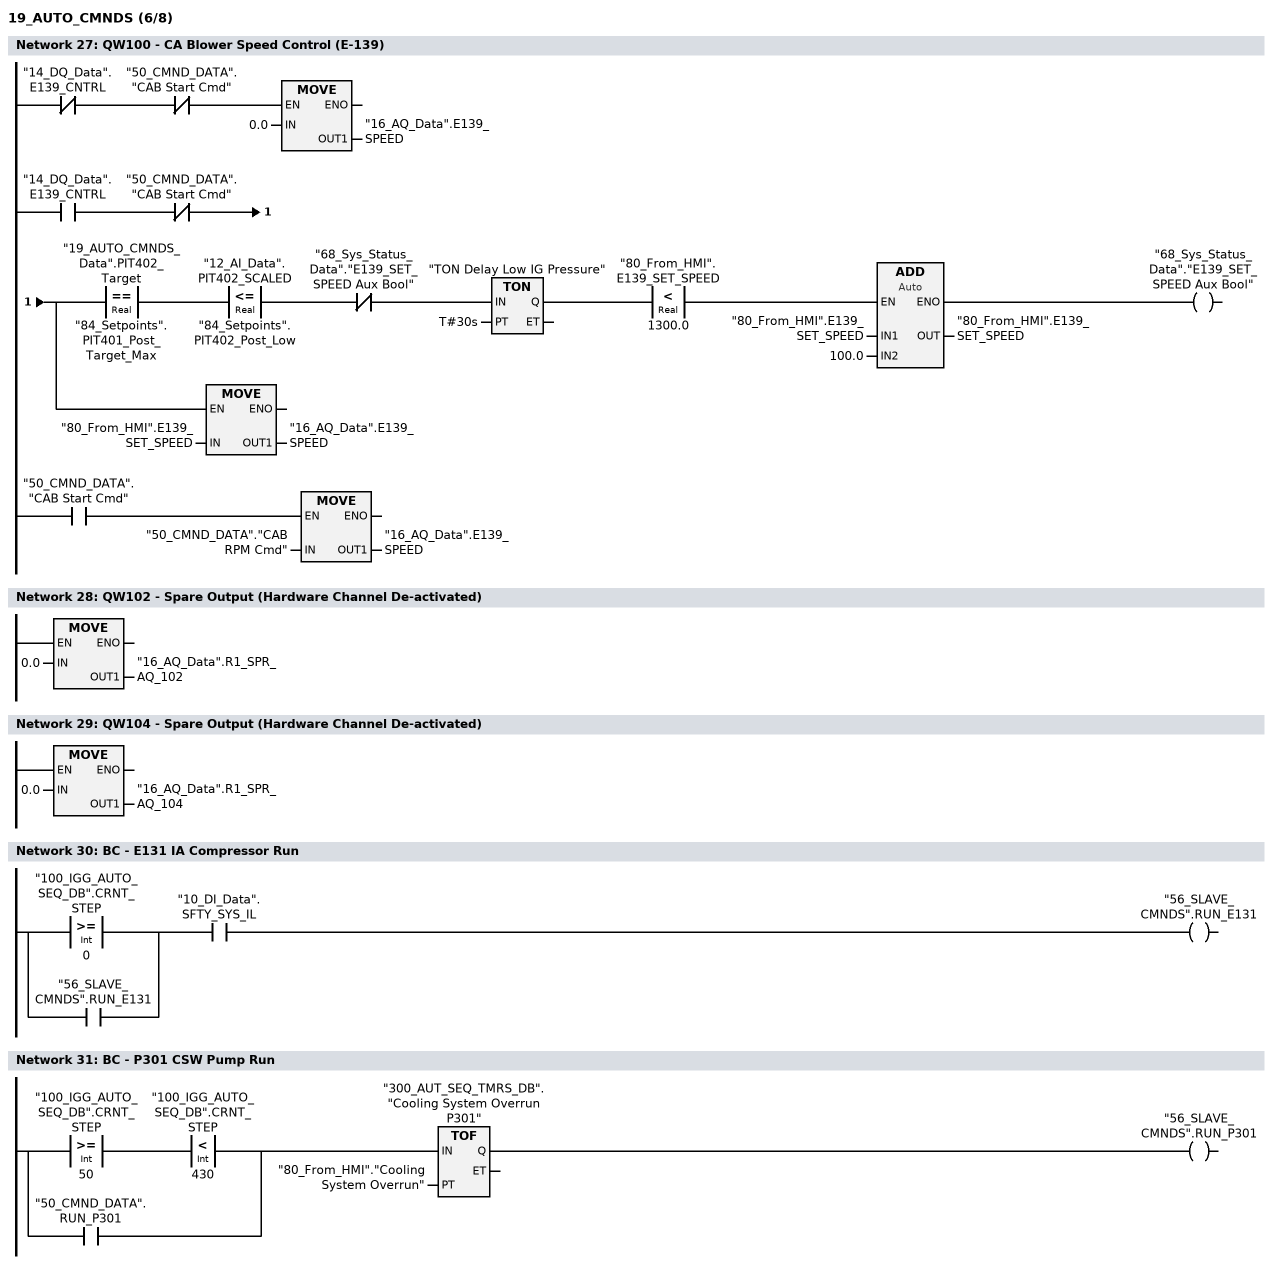
   IF NOT "14_DQ_Data".E139_CNTRL AND NOT "50_CMND_DATA"."CAB Start Cmd" THEN
       "16_AQ_Data".E139_SPEED := 0.0;
   END_IF;
   #_w1 := "14_DQ_Data".E139_CNTRL AND NOT "50_CMND_DATA"."CAB Start Cmd";
   "TON Delay Low IG Pressure".TON(IN := #_w1 AND ("19_AUTO_CMNDS_Data".PIT402_Target = "84_Setpoints".PIT401_Post_Target_Max) AND ("12_AI_Data".PIT402_SCALED <= "84_Setpoints".PIT402_Post_Low) AND NOT "68_Sys_Status_Data"."E139_SET_SPEED Aux Bool",
                           PT := T#30s);
   #_w2 := "TON Delay Low IG Pressure".Q AND ("80_From_HMI".E139_SET_SPEED < 1300.0);
   IF #_w2 THEN "80_From_HMI".E139_SET_SPEED := "80_From_HMI".E139_SET_SPEED + 100.0; END_IF;
   "68_Sys_Status_Data"."E139_SET_SPEED Aux Bool" := #_w2;
   IF #_w1 THEN "16_AQ_Data".E139_SPEED := "80_From_HMI".E139_SET_SPEED; END_IF;
   IF "50_CMND_DATA"."CAB Start Cmd" THEN "16_AQ_Data".E139_SPEED := "50_CMND_DATA"."CAB RPM Cmd"; END_IF;
END_REGION

REGION Network 28: QW102 - Spare Output (Hardware Channel De-activated)
   RUNG wire#powerrail
      Move(in := 0.0, out1 => "16_AQ_Data".R1_SPR_AQ_102)
   END_RUNG
   // the same network as SCL:
   "16_AQ_Data".R1_SPR_AQ_102 := 0.0;
END_REGION

REGION Network 29: QW104 - Spare Output (Hardware Channel De-activated)
   RUNG wire#powerrail
      Move(in := 0.0, out1 => "16_AQ_Data".R1_SPR_AQ_104)
   END_RUNG
   // the same network as SCL:
   "16_AQ_Data".R1_SPR_AQ_104 := 0.0;
END_REGION

REGION Network 30: BC - E131 IA Compressor Run
   RUNG wire#powerrail
      { S7_Templates := "SrcType := Int" } GE_Contact(in1 := "100_IGG_AUTO_SEQ_DB".CRNT_STEP, in2 := 0)
      wire#w1
      Contact( "10_DI_Data".SFTY_SYS_IL )
      Coil( "56_SLAVE_CMNDS".RUN_E131 )
   END_RUNG
   RUNG wire#powerrail
      Contact( "56_SLAVE_CMNDS".RUN_E131 )
   END_RUNG wire#w1
   // the same network as SCL:
   "56_SLAVE_CMNDS".RUN_E131 := (("100_IGG_AUTO_SEQ_DB".CRNT_STEP >= 0) OR "56_SLAVE_CMNDS".RUN_E131) AND "10_DI_Data".SFTY_SYS_IL;
END_REGION

REGION Network 31: BC - P301 CSW Pump Run
   "300_AUT_SEQ_TMRS_DB"."Cooling System Overrun P301".TOF(IN := (("100_IGG_AUTO_SEQ_DB".CRNT_STEP >= 50) AND ("100_IGG_AUTO_SEQ_DB".CRNT_STEP < 430)) OR "50_CMND_DATA".RUN_P301,
                           PT := "80_From_HMI"."Cooling System Overrun");
   "56_SLAVE_CMNDS".RUN_P301 := "300_AUT_SEQ_TMRS_DB"."Cooling System Overrun P301".Q;
END_REGION

REGION Network 32: BC - Start BC Seqence
   // Changed from 150 to5 for test
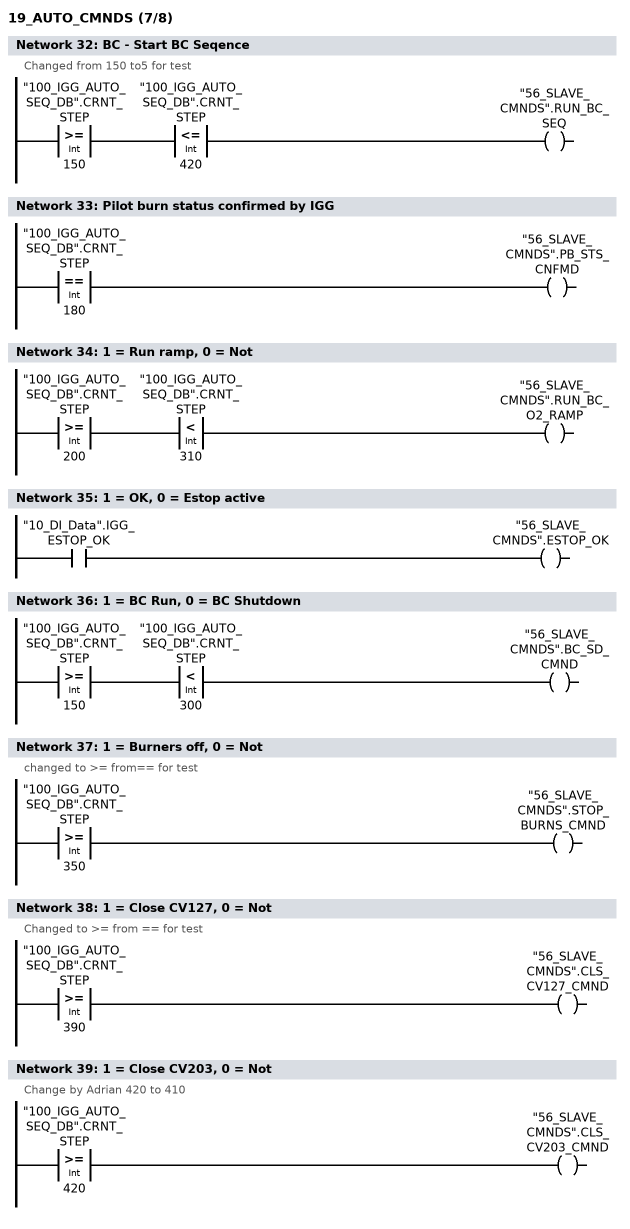
   RUNG wire#powerrail
      { S7_Templates := "SrcType := Int" } GE_Contact(in1 := "100_IGG_AUTO_SEQ_DB".CRNT_STEP, in2 := 150)
      { S7_Templates := "SrcType := Int" } LE_Contact(in1 := "100_IGG_AUTO_SEQ_DB".CRNT_STEP, in2 := 420)
      Coil( "56_SLAVE_CMNDS".RUN_BC_SEQ )
   END_RUNG
   // the same network as SCL:
   "56_SLAVE_CMNDS".RUN_BC_SEQ := ("100_IGG_AUTO_SEQ_DB".CRNT_STEP >= 150) AND ("100_IGG_AUTO_SEQ_DB".CRNT_STEP <= 420);
END_REGION

REGION Network 33: Pilot burn status confirmed by IGG
   RUNG wire#powerrail
      { S7_Templates := "SrcType := Int" } EQ_Contact(in1 := "100_IGG_AUTO_SEQ_DB".CRNT_STEP, in2 := 180)
      Coil( "56_SLAVE_CMNDS".PB_STS_CNFMD )
   END_RUNG
   // the same network as SCL:
   "56_SLAVE_CMNDS".PB_STS_CNFMD := "100_IGG_AUTO_SEQ_DB".CRNT_STEP = 180;
END_REGION

REGION Network 34: 1 = Run ramp, 0 = Not
   RUNG wire#powerrail
      { S7_Templates := "SrcType := Int" } GE_Contact(in1 := "100_IGG_AUTO_SEQ_DB".CRNT_STEP, in2 := 200)
      { S7_Templates := "SrcType := Int" } LT_Contact(in1 := "100_IGG_AUTO_SEQ_DB".CRNT_STEP, in2 := 310)
      Coil( "56_SLAVE_CMNDS".RUN_BC_O2_RAMP )
   END_RUNG
   // the same network as SCL:
   "56_SLAVE_CMNDS".RUN_BC_O2_RAMP := ("100_IGG_AUTO_SEQ_DB".CRNT_STEP >= 200) AND ("100_IGG_AUTO_SEQ_DB".CRNT_STEP < 310);
END_REGION

REGION Network 35: 1 = OK, 0 = Estop active
   RUNG wire#powerrail
      Contact( "10_DI_Data".IGG_ESTOP_OK )
      Coil( "56_SLAVE_CMNDS".ESTOP_OK )
   END_RUNG
   // the same network as SCL:
   "56_SLAVE_CMNDS".ESTOP_OK := "10_DI_Data".IGG_ESTOP_OK;
END_REGION

REGION Network 36: 1 = BC Run, 0 = BC Shutdown
   RUNG wire#powerrail
      { S7_Templates := "SrcType := Int" } GE_Contact(in1 := "100_IGG_AUTO_SEQ_DB".CRNT_STEP, in2 := 150)
      { S7_Templates := "SrcType := Int" } LT_Contact(in1 := "100_IGG_AUTO_SEQ_DB".CRNT_STEP, in2 := 300)
      Coil( "56_SLAVE_CMNDS".BC_SD_CMND )
   END_RUNG
   // the same network as SCL:
   "56_SLAVE_CMNDS".BC_SD_CMND := ("100_IGG_AUTO_SEQ_DB".CRNT_STEP >= 150) AND ("100_IGG_AUTO_SEQ_DB".CRNT_STEP < 300);
END_REGION

REGION Network 37: 1 = Burners off, 0 = Not
   // changed to >= from== for test
   RUNG wire#powerrail
      { S7_Templates := "SrcType := Int" } GE_Contact(in1 := "100_IGG_AUTO_SEQ_DB".CRNT_STEP, in2 := 350)
      Coil( "56_SLAVE_CMNDS".STOP_BURNS_CMND )
   END_RUNG
   // the same network as SCL:
   "56_SLAVE_CMNDS".STOP_BURNS_CMND := "100_IGG_AUTO_SEQ_DB".CRNT_STEP >= 350;
END_REGION

REGION Network 38: 1 = Close CV127, 0 = Not
   // Changed to >= from == for test
   RUNG wire#powerrail
      { S7_Templates := "SrcType := Int" } GE_Contact(in1 := "100_IGG_AUTO_SEQ_DB".CRNT_STEP, in2 := 390)
      Coil( "56_SLAVE_CMNDS".CLS_CV127_CMND )
   END_RUNG
   // the same network as SCL:
   "56_SLAVE_CMNDS".CLS_CV127_CMND := "100_IGG_AUTO_SEQ_DB".CRNT_STEP >= 390;
END_REGION

REGION Network 39: 1 = Close CV203, 0 = Not
   // Change by Adrian 420 to 410
   RUNG wire#powerrail
      { S7_Templates := "SrcType := Int" } GE_Contact(in1 := "100_IGG_AUTO_SEQ_DB".CRNT_STEP, in2 := 420)
      Coil( "56_SLAVE_CMNDS".CLS_CV203_CMND )
   END_RUNG
   // the same network as SCL:
   "56_SLAVE_CMNDS".CLS_CV203_CMND := "100_IGG_AUTO_SEQ_DB".CRNT_STEP >= 420;
END_REGION

REGION Network 40: 1 = Close CV111, 0 = Not
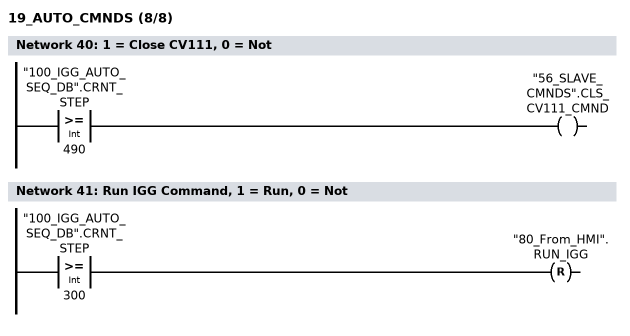
   RUNG wire#powerrail
      { S7_Templates := "SrcType := Int" } GE_Contact(in1 := "100_IGG_AUTO_SEQ_DB".CRNT_STEP, in2 := 490)
      Coil( "56_SLAVE_CMNDS".CLS_CV111_CMND )
   END_RUNG
   // the same network as SCL:
   "56_SLAVE_CMNDS".CLS_CV111_CMND := "100_IGG_AUTO_SEQ_DB".CRNT_STEP >= 490;
END_REGION

REGION Network 41: Run IGG Command, 1 = Run, 0 = Not
   RUNG wire#powerrail
      { S7_Templates := "SrcType := Int" } GE_Contact(in1 := "100_IGG_AUTO_SEQ_DB".CRNT_STEP, in2 := 300)
      R_Coil( "80_From_HMI".RUN_IGG )
   END_RUNG
   // the same network as SCL:
   IF "100_IGG_AUTO_SEQ_DB".CRNT_STEP >= 300 THEN "80_From_HMI".RUN_IGG := FALSE; END_IF;
END_REGION
END_FUNCTION

// folder: 100 - 119 Automatic Functions

FUNCTION_BLOCK "100_IGG_AUTO_SEQ"   // FB100, LAD
TITLE = Automatic Sequence
{ S7_Optimized_Access := 'TRUE' }
AUTHOR : JRS
VERSION : 0.1
// Master sequencing for automatic operation
   VAR_INPUT
      RST : Bool;   // Sequence reset
   END_VAR
   VAR_OUTPUT
      RNG : Bool;   // Sequence running
   END_VAR
   VAR
      CRNT_STEP : Int;
      STEP_001 : "500_SEQ_STEP";
      STEP_005 : "500_SEQ_STEP";
      STEP_010 : "500_SEQ_STEP";
      STEP_020 : "500_SEQ_STEP";
      STEP_030 : "500_SEQ_STEP";
      STEP_040 : "500_SEQ_STEP";
      STEP_050 : "500_SEQ_STEP";
      STEP_060 : "500_SEQ_STEP";
      STEP_070 : "500_SEQ_STEP";
      STEP_080 : "500_SEQ_STEP";
      STEP_090 : "500_SEQ_STEP";
      STEP_100 : "500_SEQ_STEP";
      STEP_110 : "500_SEQ_STEP";
      STEP_120 : "500_SEQ_STEP";
      STEP_130 : "500_SEQ_STEP";
      STEP_140 : "500_SEQ_STEP";
      STEP_150 : "500_SEQ_STEP";
      STEP_160 : "500_SEQ_STEP";
      STEP_170 : "500_SEQ_STEP";
      STEP_180 : "500_SEQ_STEP";
      STEP_190 : "500_SEQ_STEP";
      STEP_200 : "500_SEQ_STEP";
      STEP_210 : "500_SEQ_STEP";
      STEP_220 : "500_SEQ_STEP";
      STEP_300 : "500_SEQ_STEP";
      STEP_310 : "500_SEQ_STEP";
      STEP_320 : "500_SEQ_STEP";
      STEP_330 : "500_SEQ_STEP";
      STEP_340 : "500_SEQ_STEP";
      STEP_350 : "500_SEQ_STEP";
      STEP_360 : "500_SEQ_STEP";
      STEP_370 : "500_SEQ_STEP";
      STEP_380 : "500_SEQ_STEP";
      STEP_390 : "500_SEQ_STEP";
      STEP_400 : "500_SEQ_STEP";
      STEP_410 : "500_SEQ_STEP";
      STEP_420 : "500_SEQ_STEP";
      STEP_430 : "500_SEQ_STEP";
      STEP_440 : "500_SEQ_STEP";
      STEP_450 : "500_SEQ_STEP";
      STEP_460 : "500_SEQ_STEP";
      STEP_470 : "500_SEQ_STEP";
      STEP_480 : "500_SEQ_STEP";
      STEP_490 : "500_SEQ_STEP";
      STEP_500 : "500_SEQ_STEP";
      Aux : Struct
         Aux1 : Bool;
         Aux2 : Bool;
         Aux3 : Bool;
      END_STRUCT;
      IEC_Timer_0_Instance : TP_TIME;
   END_VAR
   VAR_TEMP   // added for the SCL form of the ladder/FBD networks
      _w1 : Bool;
      _w2 : Bool;
   END_VAR
BEGIN

REGION Network 1: Auto Initiated or Reset = Set Step to 0
   // Going into automatic or sequence reset resets the sequence
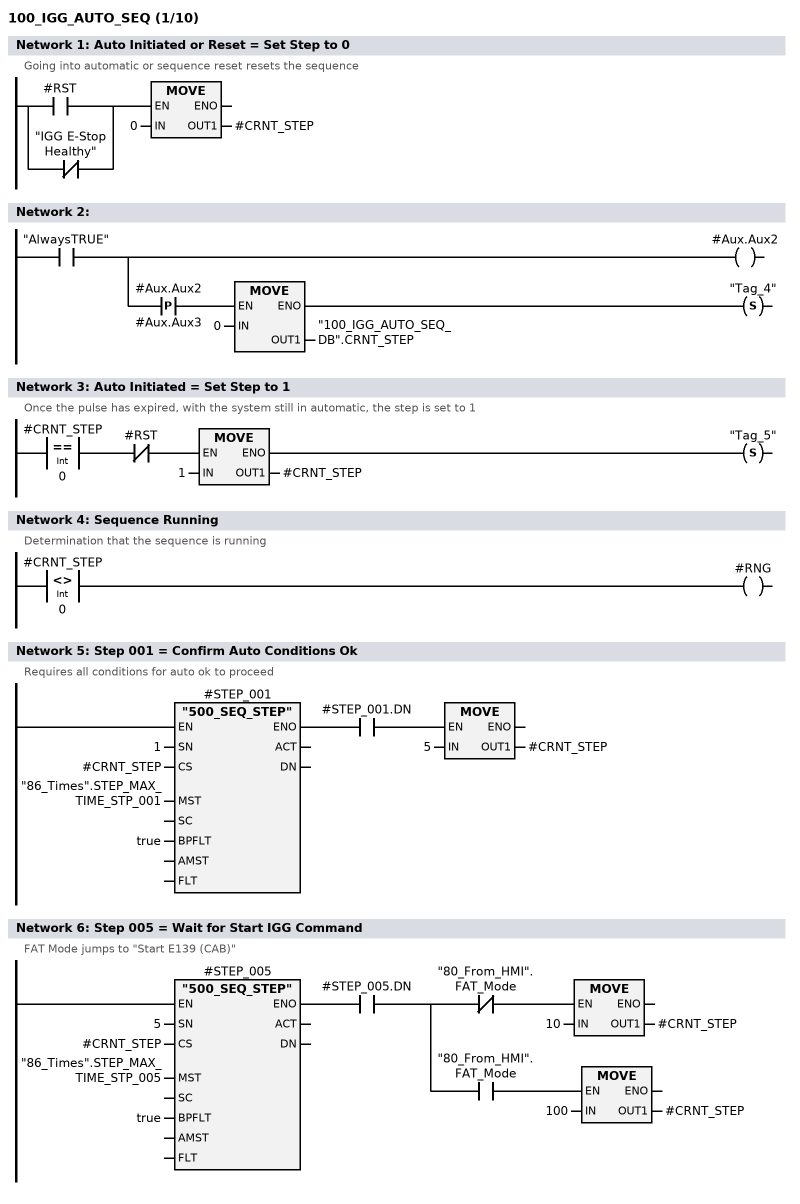
   RUNG wire#powerrail
      Contact( #RST )
      wire#w1
      Move(in := 0, out1 => #CRNT_STEP)
   END_RUNG
   RUNG wire#powerrail
      I_Contact( "IGG E-Stop Healthy" )
   END_RUNG wire#w1
   // the same network as SCL:
   IF #RST OR NOT "IGG E-Stop Healthy" THEN #CRNT_STEP := 0; END_IF;
END_REGION

REGION Network 2
   RUNG wire#powerrail
      Contact( "AlwaysTRUE" )
      wire#w1
      Coil( #Aux.Aux2 )
   END_RUNG
   RUNG wire#w1
      P_Contact(operand := #Aux.Aux2, bit := #Aux.Aux3)
      Move(in := 0, out1 => "100_IGG_AUTO_SEQ_DB".CRNT_STEP)
      S_Coil( "Tag_4" )
   END_RUNG
   // the same network as SCL:
   #Aux.Aux2 := "AlwaysTRUE";
   #_w1 := "AlwaysTRUE" AND #Aux.Aux2 AND NOT #Aux.Aux3;   // rising edge of #Aux.Aux2
   #Aux.Aux3 := #Aux.Aux2;
   IF #_w1 THEN
       "100_IGG_AUTO_SEQ_DB".CRNT_STEP := 0;
       "Tag_4" := TRUE;
   END_IF;
END_REGION

REGION Network 3: Auto Initiated = Set Step to 1
   // Once the pulse has expired, with the system still in automatic, the step is set to 1
   RUNG wire#powerrail
      { S7_Templates := "SrcType := Int" } EQ_Contact(in1 := #CRNT_STEP, in2 := 0)
      I_Contact( #RST )
      Move(in := 1, out1 => #CRNT_STEP)
      S_Coil( "Tag_5" )
   END_RUNG
   // the same network as SCL:
   #_w1 := (#CRNT_STEP = 0) AND NOT #RST;
   IF #_w1 THEN
       #CRNT_STEP := 1;
       "Tag_5" := TRUE;
   END_IF;
END_REGION

REGION Network 4: Sequence Running
   // Determination that the sequence is running
   RUNG wire#powerrail
      { S7_Templates := "SrcType := Int" } NE_Contact(in1 := #CRNT_STEP, in2 := 0)
      Coil( #RNG )
   END_RUNG
   // the same network as SCL:
   #RNG := #CRNT_STEP <> 0;
END_REGION

REGION Network 5: Step 001 = Confirm Auto Conditions Ok
   // Requires all conditions for auto ok to proceed
   RUNG wire#powerrail
      #STEP_001(SN := 1, CS := #CRNT_STEP, MST := "86_Times".STEP_MAX_TIME_STP_001, SC :=, BPFLT := true, AMST :=, FLT :=, ACT =>, DN =>)
      Contact( #STEP_001.DN )
      Move(in := 5, out1 => #CRNT_STEP)
   END_RUNG
   // the same network as SCL:
   #STEP_001(SN := 1, CS := #CRNT_STEP, MST := "86_Times".STEP_MAX_TIME_STP_001, BPFLT := true, ENO => #_w1);   // "500_SEQ_STEP"
   IF #_w1 AND #STEP_001.DN THEN #CRNT_STEP := 5; END_IF;
END_REGION

REGION Network 6: Step 005 = Wait for Start IGG Command
   // FAT Mode jumps to "Start E139 (CAB)"
   RUNG wire#powerrail
      #STEP_005(SN := 5, CS := #CRNT_STEP, MST := "86_Times".STEP_MAX_TIME_STP_005, SC :=, BPFLT := true, AMST :=, FLT :=, ACT =>, DN =>)
      Contact( #STEP_005.DN )
      wire#w1
      I_Contact( "80_From_HMI".FAT_Mode )
      Move(in := 10, out1 => #CRNT_STEP)
   END_RUNG
   RUNG wire#w1
      Contact( "80_From_HMI".FAT_Mode )
      Move(in := 100, out1 => #CRNT_STEP)
   END_RUNG
   // the same network as SCL:
   #STEP_005(SN := 5, CS := #CRNT_STEP, MST := "86_Times".STEP_MAX_TIME_STP_005, BPFLT := true, ENO => #_w1);   // "500_SEQ_STEP"
   #_w2 := #_w1 AND #STEP_005.DN;
   IF #_w2 AND NOT "80_From_HMI".FAT_Mode THEN #CRNT_STEP := 10; END_IF;
   IF #_w2 AND "80_From_HMI".FAT_Mode THEN #CRNT_STEP := 100; END_IF;
END_REGION

REGION Network 7: Step 010 = Start E131 (IA Compressor)
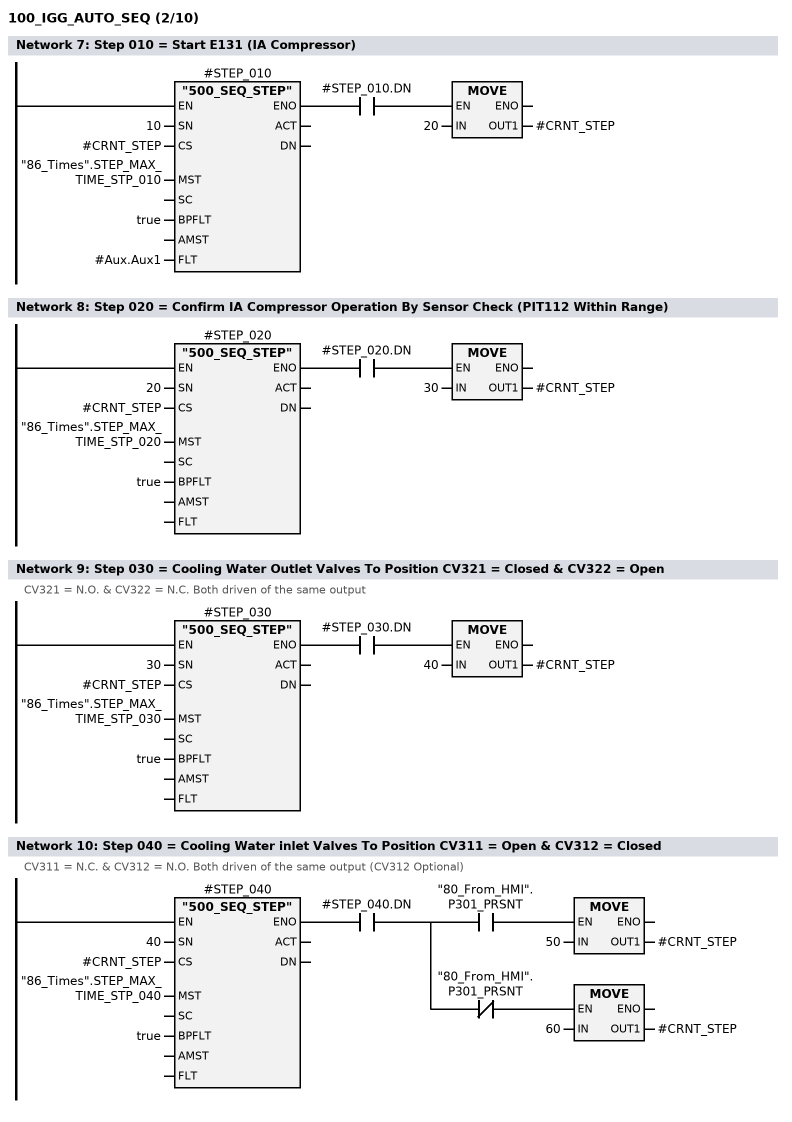
   RUNG wire#powerrail
      #STEP_010(SN := 10, CS := #CRNT_STEP, MST := "86_Times".STEP_MAX_TIME_STP_010, SC :=, BPFLT := true, AMST :=, FLT := #Aux.Aux1, ACT =>, DN =>)
      Contact( #STEP_010.DN )
      Move(in := 20, out1 => #CRNT_STEP)
   END_RUNG
   // the same network as SCL:
   #STEP_010(SN := 10,   // "500_SEQ_STEP"
             CS := #CRNT_STEP,
             MST := "86_Times".STEP_MAX_TIME_STP_010,
             BPFLT := true,
             FLT := #Aux.Aux1,
             ENO => #_w1);
   IF #_w1 AND #STEP_010.DN THEN #CRNT_STEP := 20; END_IF;
END_REGION

REGION Network 8: Step 020 = Confirm IA Compressor Operation By Sensor Check (PIT112 Within Range)
   RUNG wire#powerrail
      #STEP_020(SN := 20, CS := #CRNT_STEP, MST := "86_Times".STEP_MAX_TIME_STP_020, SC :=, BPFLT := true, AMST :=, FLT :=, ACT =>, DN =>)
      Contact( #STEP_020.DN )
      Move(in := 30, out1 => #CRNT_STEP)
   END_RUNG
   // the same network as SCL:
   #STEP_020(SN := 20, CS := #CRNT_STEP, MST := "86_Times".STEP_MAX_TIME_STP_020, BPFLT := true, ENO => #_w1);   // "500_SEQ_STEP"
   IF #_w1 AND #STEP_020.DN THEN #CRNT_STEP := 30; END_IF;
END_REGION

REGION Network 9: Step 030 = Cooling Water Outlet Valves To Position CV321 = Closed & CV322 = Open
   // CV321 = N.O. & CV322 = N.C. Both driven of the same output
   RUNG wire#powerrail
      #STEP_030(SN := 30, CS := #CRNT_STEP, MST := "86_Times".STEP_MAX_TIME_STP_030, SC :=, BPFLT := true, AMST :=, FLT :=, ACT =>, DN =>)
      Contact( #STEP_030.DN )
      Move(in := 40, out1 => #CRNT_STEP)
   END_RUNG
   // the same network as SCL:
   #STEP_030(SN := 30, CS := #CRNT_STEP, MST := "86_Times".STEP_MAX_TIME_STP_030, BPFLT := true, ENO => #_w1);   // "500_SEQ_STEP"
   IF #_w1 AND #STEP_030.DN THEN #CRNT_STEP := 40; END_IF;
END_REGION

REGION Network 10: Step 040 = Cooling Water inlet Valves To Position CV311 = Open & CV312 = Closed
   // CV311 = N.C. & CV312 = N.O. Both driven of the same output (CV312 Optional)
   RUNG wire#powerrail
      #STEP_040(SN := 40, CS := #CRNT_STEP, MST := "86_Times".STEP_MAX_TIME_STP_040, SC :=, BPFLT := true, AMST :=, FLT :=, ACT =>, DN =>)
      Contact( #STEP_040.DN )
      wire#w1
      Contact( "80_From_HMI".P301_PRSNT )
      Move(in := 50, out1 => #CRNT_STEP)
   END_RUNG
   RUNG wire#w1
      I_Contact( "80_From_HMI".P301_PRSNT )
      Move(in := 60, out1 => #CRNT_STEP)
   END_RUNG
   // the same network as SCL:
   #STEP_040(SN := 40, CS := #CRNT_STEP, MST := "86_Times".STEP_MAX_TIME_STP_040, BPFLT := true, ENO => #_w1);   // "500_SEQ_STEP"
   #_w2 := #_w1 AND #STEP_040.DN;
   IF #_w2 AND "80_From_HMI".P301_PRSNT THEN #CRNT_STEP := 50; END_IF;
   IF #_w2 AND NOT "80_From_HMI".P301_PRSNT THEN #CRNT_STEP := 60; END_IF;
END_REGION

REGION Network 11: Step 050 = Start P301 (CSW Pump)
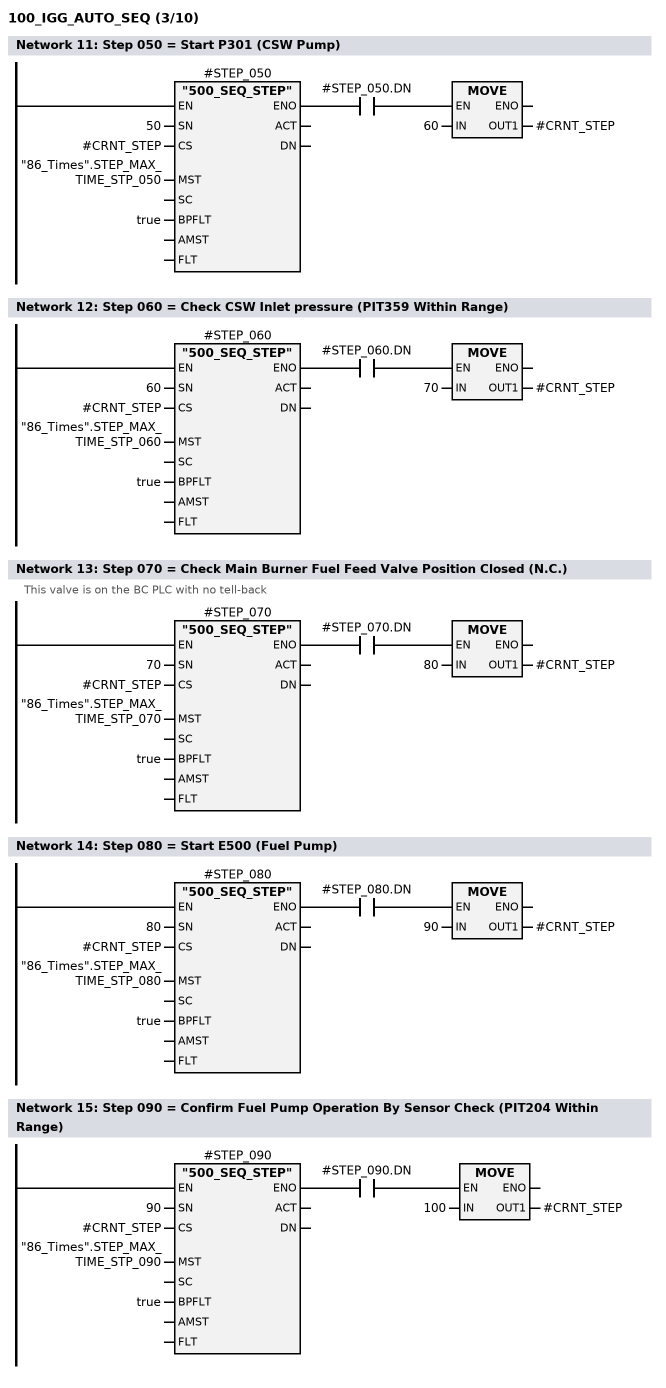
   RUNG wire#powerrail
      #STEP_050(SN := 50, CS := #CRNT_STEP, MST := "86_Times".STEP_MAX_TIME_STP_050, SC :=, BPFLT := true, AMST :=, FLT :=, ACT =>, DN =>)
      Contact( #STEP_050.DN )
      Move(in := 60, out1 => #CRNT_STEP)
   END_RUNG
   // the same network as SCL:
   #STEP_050(SN := 50, CS := #CRNT_STEP, MST := "86_Times".STEP_MAX_TIME_STP_050, BPFLT := true, ENO => #_w1);   // "500_SEQ_STEP"
   IF #_w1 AND #STEP_050.DN THEN #CRNT_STEP := 60; END_IF;
END_REGION

REGION Network 12: Step 060 = Check CSW Inlet pressure (PIT359 Within Range)
   RUNG wire#powerrail
      #STEP_060(SN := 60, CS := #CRNT_STEP, MST := "86_Times".STEP_MAX_TIME_STP_060, SC :=, BPFLT := true, AMST :=, FLT :=, ACT =>, DN =>)
      Contact( #STEP_060.DN )
      Move(in := 70, out1 => #CRNT_STEP)
   END_RUNG
   // the same network as SCL:
   #STEP_060(SN := 60, CS := #CRNT_STEP, MST := "86_Times".STEP_MAX_TIME_STP_060, BPFLT := true, ENO => #_w1);   // "500_SEQ_STEP"
   IF #_w1 AND #STEP_060.DN THEN #CRNT_STEP := 70; END_IF;
END_REGION

REGION Network 13: Step 070 = Check Main Burner Fuel Feed Valve Position Closed (N.C.)
   // This valve is on the BC PLC with no tell-back
   RUNG wire#powerrail
      #STEP_070(SN := 70, CS := #CRNT_STEP, MST := "86_Times".STEP_MAX_TIME_STP_070, SC :=, BPFLT := true, AMST :=, FLT :=, ACT =>, DN =>)
      Contact( #STEP_070.DN )
      Move(in := 80, out1 => #CRNT_STEP)
   END_RUNG
   // the same network as SCL:
   #STEP_070(SN := 70, CS := #CRNT_STEP, MST := "86_Times".STEP_MAX_TIME_STP_070, BPFLT := true, ENO => #_w1);   // "500_SEQ_STEP"
   IF #_w1 AND #STEP_070.DN THEN #CRNT_STEP := 80; END_IF;
END_REGION

REGION Network 14: Step 080 = Start E500 (Fuel Pump)
   RUNG wire#powerrail
      #STEP_080(SN := 80, CS := #CRNT_STEP, MST := "86_Times".STEP_MAX_TIME_STP_080, SC :=, BPFLT := true, AMST :=, FLT :=, ACT =>, DN =>)
      Contact( #STEP_080.DN )
      Move(in := 90, out1 => #CRNT_STEP)
   END_RUNG
   // the same network as SCL:
   #STEP_080(SN := 80, CS := #CRNT_STEP, MST := "86_Times".STEP_MAX_TIME_STP_080, BPFLT := true, ENO => #_w1);   // "500_SEQ_STEP"
   IF #_w1 AND #STEP_080.DN THEN #CRNT_STEP := 90; END_IF;
END_REGION

REGION Network 15: Step 090 = Confirm Fuel Pump Operation By Sensor Check (PIT204 Within Range)
   RUNG wire#powerrail
      #STEP_090(SN := 90, CS := #CRNT_STEP, MST := "86_Times".STEP_MAX_TIME_STP_090, SC :=, BPFLT := true, AMST :=, FLT :=, ACT =>, DN =>)
      Contact( #STEP_090.DN )
      Move(in := 100, out1 => #CRNT_STEP)
   END_RUNG
   // the same network as SCL:
   #STEP_090(SN := 90, CS := #CRNT_STEP, MST := "86_Times".STEP_MAX_TIME_STP_090, BPFLT := true, ENO => #_w1);   // "500_SEQ_STEP"
   IF #_w1 AND #STEP_090.DN THEN #CRNT_STEP := 100; END_IF;
END_REGION

REGION Network 16: Step 100 = Start E139 (CAB)
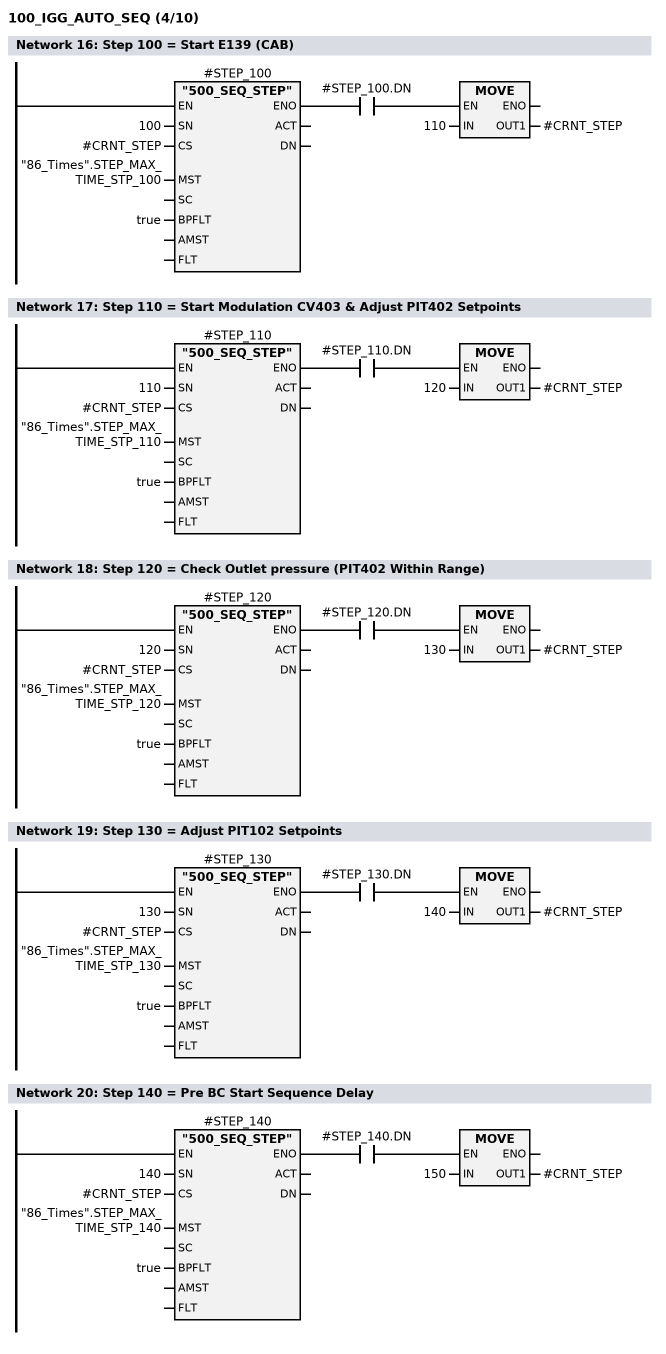
   RUNG wire#powerrail
      #STEP_100(SN := 100, CS := #CRNT_STEP, MST := "86_Times".STEP_MAX_TIME_STP_100, SC :=, BPFLT := true, AMST :=, FLT :=, ACT =>, DN =>)
      Contact( #STEP_100.DN )
      Move(in := 110, out1 => #CRNT_STEP)
   END_RUNG
   // the same network as SCL:
   #STEP_100(SN := 100, CS := #CRNT_STEP, MST := "86_Times".STEP_MAX_TIME_STP_100, BPFLT := true, ENO => #_w1);   // "500_SEQ_STEP"
   IF #_w1 AND #STEP_100.DN THEN #CRNT_STEP := 110; END_IF;
END_REGION

REGION Network 17: Step 110 = Start Modulation CV403 & Adjust PIT402 Setpoints
   RUNG wire#powerrail
      #STEP_110(SN := 110, CS := #CRNT_STEP, MST := "86_Times".STEP_MAX_TIME_STP_110, SC :=, BPFLT := true, AMST :=, FLT :=, ACT =>, DN =>)
      Contact( #STEP_110.DN )
      Move(in := 120, out1 => #CRNT_STEP)
   END_RUNG
   // the same network as SCL:
   #STEP_110(SN := 110, CS := #CRNT_STEP, MST := "86_Times".STEP_MAX_TIME_STP_110, BPFLT := true, ENO => #_w1);   // "500_SEQ_STEP"
   IF #_w1 AND #STEP_110.DN THEN #CRNT_STEP := 120; END_IF;
END_REGION

REGION Network 18: Step 120 = Check Outlet pressure (PIT402 Within Range)
   RUNG wire#powerrail
      #STEP_120(SN := 120, CS := #CRNT_STEP, MST := "86_Times".STEP_MAX_TIME_STP_120, SC :=, BPFLT := true, AMST :=, FLT :=, ACT =>, DN =>)
      Contact( #STEP_120.DN )
      Move(in := 130, out1 => #CRNT_STEP)
   END_RUNG
   // the same network as SCL:
   #STEP_120(SN := 120, CS := #CRNT_STEP, MST := "86_Times".STEP_MAX_TIME_STP_120, BPFLT := true, ENO => #_w1);   // "500_SEQ_STEP"
   IF #_w1 AND #STEP_120.DN THEN #CRNT_STEP := 130; END_IF;
END_REGION

REGION Network 19: Step 130 = Adjust PIT102 Setpoints
   RUNG wire#powerrail
      #STEP_130(SN := 130, CS := #CRNT_STEP, MST := "86_Times".STEP_MAX_TIME_STP_130, SC :=, BPFLT := true, AMST :=, FLT :=, ACT =>, DN =>)
      Contact( #STEP_130.DN )
      Move(in := 140, out1 => #CRNT_STEP)
   END_RUNG
   // the same network as SCL:
   #STEP_130(SN := 130, CS := #CRNT_STEP, MST := "86_Times".STEP_MAX_TIME_STP_130, BPFLT := true, ENO => #_w1);   // "500_SEQ_STEP"
   IF #_w1 AND #STEP_130.DN THEN #CRNT_STEP := 140; END_IF;
END_REGION

REGION Network 20: Step 140 = Pre BC Start Sequence Delay
   RUNG wire#powerrail
      #STEP_140(SN := 140, CS := #CRNT_STEP, MST := "86_Times".STEP_MAX_TIME_STP_140, SC :=, BPFLT := true, AMST :=, FLT :=, ACT =>, DN =>)
      Contact( #STEP_140.DN )
      Move(in := 150, out1 => #CRNT_STEP)
   END_RUNG
   // the same network as SCL:
   #STEP_140(SN := 140, CS := #CRNT_STEP, MST := "86_Times".STEP_MAX_TIME_STP_140, BPFLT := true, ENO => #_w1);   // "500_SEQ_STEP"
   IF #_w1 AND #STEP_140.DN THEN #CRNT_STEP := 150; END_IF;
END_REGION

REGION Network 21: Step 150 = BC Start Command
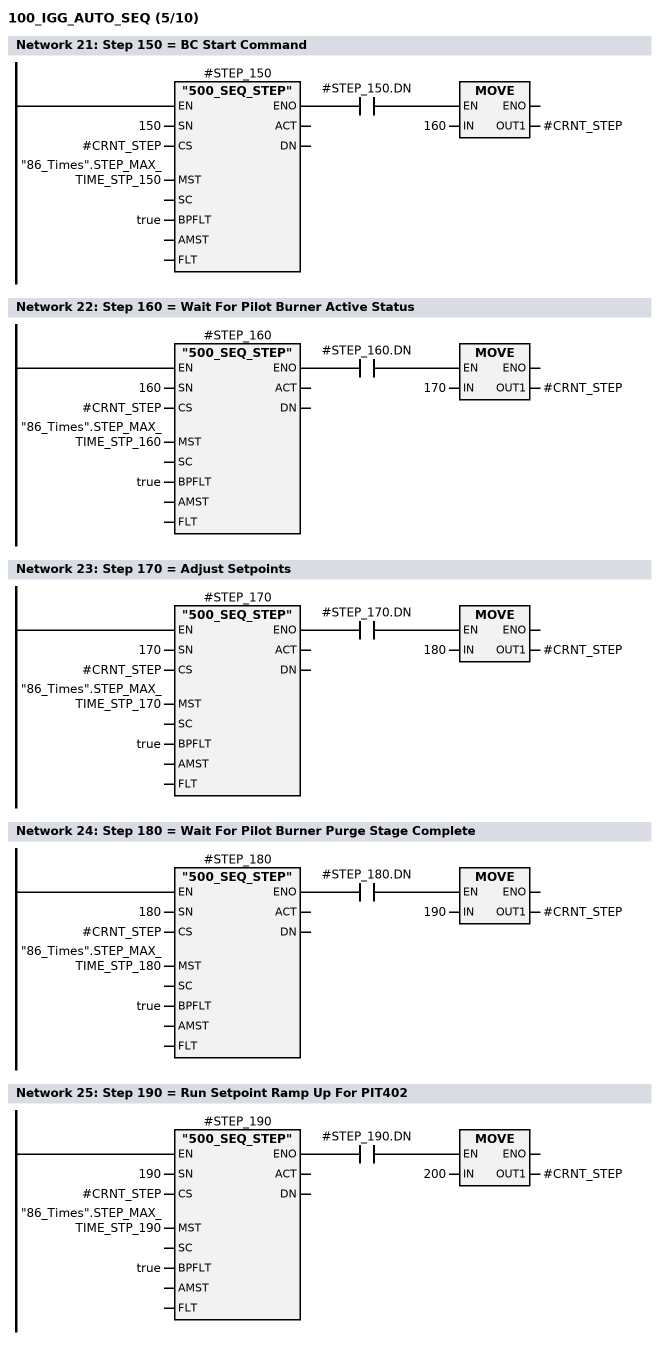
   RUNG wire#powerrail
      #STEP_150(SN := 150, CS := #CRNT_STEP, MST := "86_Times".STEP_MAX_TIME_STP_150, SC :=, BPFLT := true, AMST :=, FLT :=, ACT =>, DN =>)
      Contact( #STEP_150.DN )
      Move(in := 160, out1 => #CRNT_STEP)
   END_RUNG
   // the same network as SCL:
   #STEP_150(SN := 150, CS := #CRNT_STEP, MST := "86_Times".STEP_MAX_TIME_STP_150, BPFLT := true, ENO => #_w1);   // "500_SEQ_STEP"
   IF #_w1 AND #STEP_150.DN THEN #CRNT_STEP := 160; END_IF;
END_REGION

REGION Network 22: Step 160 = Wait For Pilot Burner Active Status
   RUNG wire#powerrail
      #STEP_160(SN := 160, CS := #CRNT_STEP, MST := "86_Times".STEP_MAX_TIME_STP_160, SC :=, BPFLT := true, AMST :=, FLT :=, ACT =>, DN =>)
      Contact( #STEP_160.DN )
      Move(in := 170, out1 => #CRNT_STEP)
   END_RUNG
   // the same network as SCL:
   #STEP_160(SN := 160, CS := #CRNT_STEP, MST := "86_Times".STEP_MAX_TIME_STP_160, BPFLT := true, ENO => #_w1);   // "500_SEQ_STEP"
   IF #_w1 AND #STEP_160.DN THEN #CRNT_STEP := 170; END_IF;
END_REGION

REGION Network 23: Step 170 = Adjust Setpoints
   RUNG wire#powerrail
      #STEP_170(SN := 170, CS := #CRNT_STEP, MST := "86_Times".STEP_MAX_TIME_STP_170, SC :=, BPFLT := true, AMST :=, FLT :=, ACT =>, DN =>)
      Contact( #STEP_170.DN )
      Move(in := 180, out1 => #CRNT_STEP)
   END_RUNG
   // the same network as SCL:
   #STEP_170(SN := 170, CS := #CRNT_STEP, MST := "86_Times".STEP_MAX_TIME_STP_170, BPFLT := true, ENO => #_w1);   // "500_SEQ_STEP"
   IF #_w1 AND #STEP_170.DN THEN #CRNT_STEP := 180; END_IF;
END_REGION

REGION Network 24: Step 180 = Wait For Pilot Burner Purge Stage Complete
   RUNG wire#powerrail
      #STEP_180(SN := 180, CS := #CRNT_STEP, MST := "86_Times".STEP_MAX_TIME_STP_180, SC :=, BPFLT := true, AMST :=, FLT :=, ACT =>, DN =>)
      Contact( #STEP_180.DN )
      Move(in := 190, out1 => #CRNT_STEP)
   END_RUNG
   // the same network as SCL:
   #STEP_180(SN := 180, CS := #CRNT_STEP, MST := "86_Times".STEP_MAX_TIME_STP_180, BPFLT := true, ENO => #_w1);   // "500_SEQ_STEP"
   IF #_w1 AND #STEP_180.DN THEN #CRNT_STEP := 190; END_IF;
END_REGION

REGION Network 25: Step 190 = Run Setpoint Ramp Up For PIT402
   RUNG wire#powerrail
      #STEP_190(SN := 190, CS := #CRNT_STEP, MST := "86_Times".STEP_MAX_TIME_STP_190, SC :=, BPFLT := true, AMST :=, FLT :=, ACT =>, DN =>)
      Contact( #STEP_190.DN )
      Move(in := 200, out1 => #CRNT_STEP)
   END_RUNG
   // the same network as SCL:
   #STEP_190(SN := 190, CS := #CRNT_STEP, MST := "86_Times".STEP_MAX_TIME_STP_190, BPFLT := true, ENO => #_w1);   // "500_SEQ_STEP"
   IF #_w1 AND #STEP_190.DN THEN #CRNT_STEP := 200; END_IF;
END_REGION

REGION Network 26: Step 200 = BC Ramp O2 Command